// TIA Portal project "XSFW_TIA31001_B0_V15.1" (V15.1) (continued)
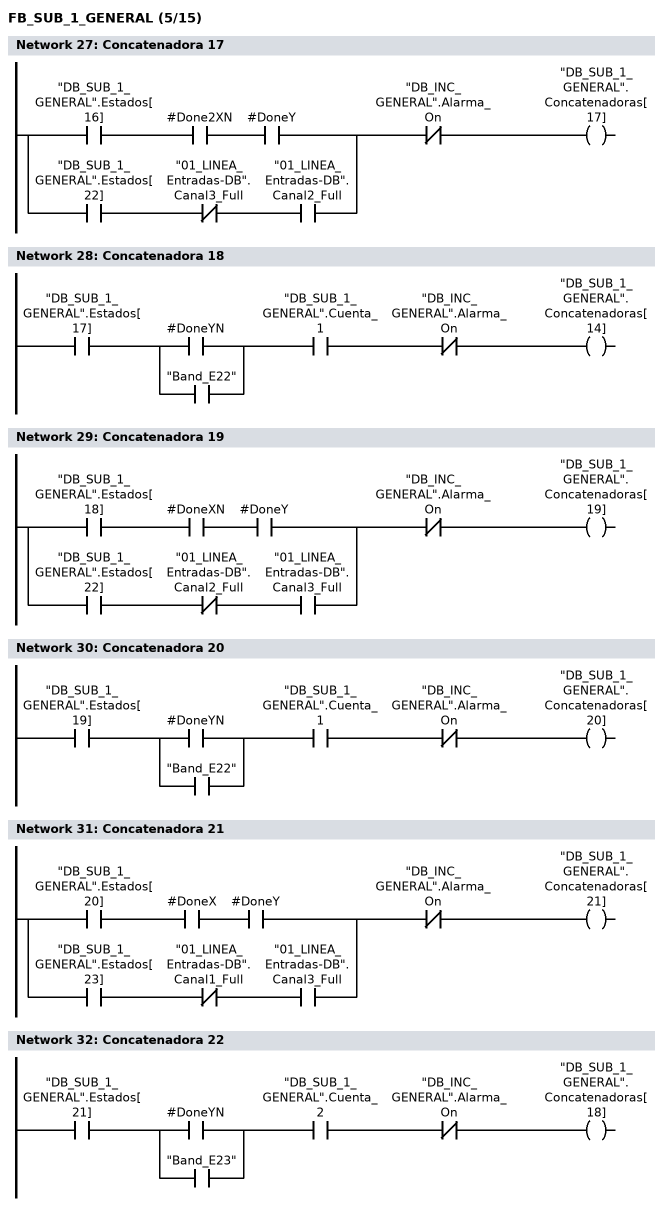
   RUNG wire#powerrail
      Contact( "DB_SUB_1_GENERAL".Estados[16] )
      Contact( #Done2XN )
      Contact( #DoneY )
      wire#w1
      I_Contact( "DB_INC_GENERAL".Alarma_On )
      Coil( "DB_SUB_1_GENERAL".Concatenadoras[17] )
   END_RUNG
   RUNG wire#powerrail
      Contact( "DB_SUB_1_GENERAL".Estados[22] )
      I_Contact( "01_LINEA_Entradas-DB".Canal3_Full )
      Contact( "01_LINEA_Entradas-DB".Canal2_Full )
   END_RUNG wire#w1
   // the same network as SCL:
   "DB_SUB_1_GENERAL".Concatenadoras[17] := (("DB_SUB_1_GENERAL".Estados[16] AND #Done2XN AND #DoneY) OR ("DB_SUB_1_GENERAL".Estados[22] AND NOT "01_LINEA_Entradas-DB".Canal3_Full AND "01_LINEA_Entradas-DB".Canal2_Full)) AND NOT "DB_INC_GENERAL".Alarma_On;
END_REGION

REGION Network 28: Concatenadora 18
   RUNG wire#powerrail
      Contact( "DB_SUB_1_GENERAL".Estados[17] )
      wire#w1
      Contact( #DoneYN )
      wire#w2
      Contact( "DB_SUB_1_GENERAL".Cuenta_1 )
      I_Contact( "DB_INC_GENERAL".Alarma_On )
      Coil( "DB_SUB_1_GENERAL".Concatenadoras[14] )
   END_RUNG
   RUNG wire#w1
      Contact( "Band_E22" )
   END_RUNG wire#w2
   // the same network as SCL:
   "DB_SUB_1_GENERAL".Concatenadoras[14] := "DB_SUB_1_GENERAL".Estados[17] AND (#DoneYN OR "Band_E22") AND "DB_SUB_1_GENERAL".Cuenta_1 AND NOT "DB_INC_GENERAL".Alarma_On;
END_REGION

REGION Network 29: Concatenadora 19
   RUNG wire#powerrail
      Contact( "DB_SUB_1_GENERAL".Estados[18] )
      Contact( #DoneXN )
      Contact( #DoneY )
      wire#w1
      I_Contact( "DB_INC_GENERAL".Alarma_On )
      Coil( "DB_SUB_1_GENERAL".Concatenadoras[19] )
   END_RUNG
   RUNG wire#powerrail
      Contact( "DB_SUB_1_GENERAL".Estados[22] )
      I_Contact( "01_LINEA_Entradas-DB".Canal2_Full )
      Contact( "01_LINEA_Entradas-DB".Canal3_Full )
   END_RUNG wire#w1
   // the same network as SCL:
   "DB_SUB_1_GENERAL".Concatenadoras[19] := (("DB_SUB_1_GENERAL".Estados[18] AND #DoneXN AND #DoneY) OR ("DB_SUB_1_GENERAL".Estados[22] AND NOT "01_LINEA_Entradas-DB".Canal2_Full AND "01_LINEA_Entradas-DB".Canal3_Full)) AND NOT "DB_INC_GENERAL".Alarma_On;
END_REGION

REGION Network 30: Concatenadora 20
   RUNG wire#powerrail
      Contact( "DB_SUB_1_GENERAL".Estados[19] )
      wire#w1
      Contact( #DoneYN )
      wire#w2
      Contact( "DB_SUB_1_GENERAL".Cuenta_1 )
      I_Contact( "DB_INC_GENERAL".Alarma_On )
      Coil( "DB_SUB_1_GENERAL".Concatenadoras[20] )
   END_RUNG
   RUNG wire#w1
      Contact( "Band_E22" )
   END_RUNG wire#w2
   // the same network as SCL:
   "DB_SUB_1_GENERAL".Concatenadoras[20] := "DB_SUB_1_GENERAL".Estados[19] AND (#DoneYN OR "Band_E22") AND "DB_SUB_1_GENERAL".Cuenta_1 AND NOT "DB_INC_GENERAL".Alarma_On;
END_REGION

REGION Network 31: Concatenadora 21
   RUNG wire#powerrail
      Contact( "DB_SUB_1_GENERAL".Estados[20] )
      Contact( #DoneX )
      Contact( #DoneY )
      wire#w1
      I_Contact( "DB_INC_GENERAL".Alarma_On )
      Coil( "DB_SUB_1_GENERAL".Concatenadoras[21] )
   END_RUNG
   RUNG wire#powerrail
      Contact( "DB_SUB_1_GENERAL".Estados[23] )
      I_Contact( "01_LINEA_Entradas-DB".Canal1_Full )
      Contact( "01_LINEA_Entradas-DB".Canal3_Full )
   END_RUNG wire#w1
   // the same network as SCL:
   "DB_SUB_1_GENERAL".Concatenadoras[21] := (("DB_SUB_1_GENERAL".Estados[20] AND #DoneX AND #DoneY) OR ("DB_SUB_1_GENERAL".Estados[23] AND NOT "01_LINEA_Entradas-DB".Canal1_Full AND "01_LINEA_Entradas-DB".Canal3_Full)) AND NOT "DB_INC_GENERAL".Alarma_On;
END_REGION

REGION Network 32: Concatenadora 22
   RUNG wire#powerrail
      Contact( "DB_SUB_1_GENERAL".Estados[21] )
      wire#w1
      Contact( #DoneYN )
      wire#w2
      Contact( "DB_SUB_1_GENERAL".Cuenta_2 )
      I_Contact( "DB_INC_GENERAL".Alarma_On )
      Coil( "DB_SUB_1_GENERAL".Concatenadoras[18] )
   END_RUNG
   RUNG wire#w1
      Contact( "Band_E23" )
   END_RUNG wire#w2
   // the same network as SCL:
   "DB_SUB_1_GENERAL".Concatenadoras[18] := "DB_SUB_1_GENERAL".Estados[21] AND (#DoneYN OR "Band_E23") AND "DB_SUB_1_GENERAL".Cuenta_2 AND NOT "DB_INC_GENERAL".Alarma_On;
END_REGION

REGION Network 33: Prioritaria 0
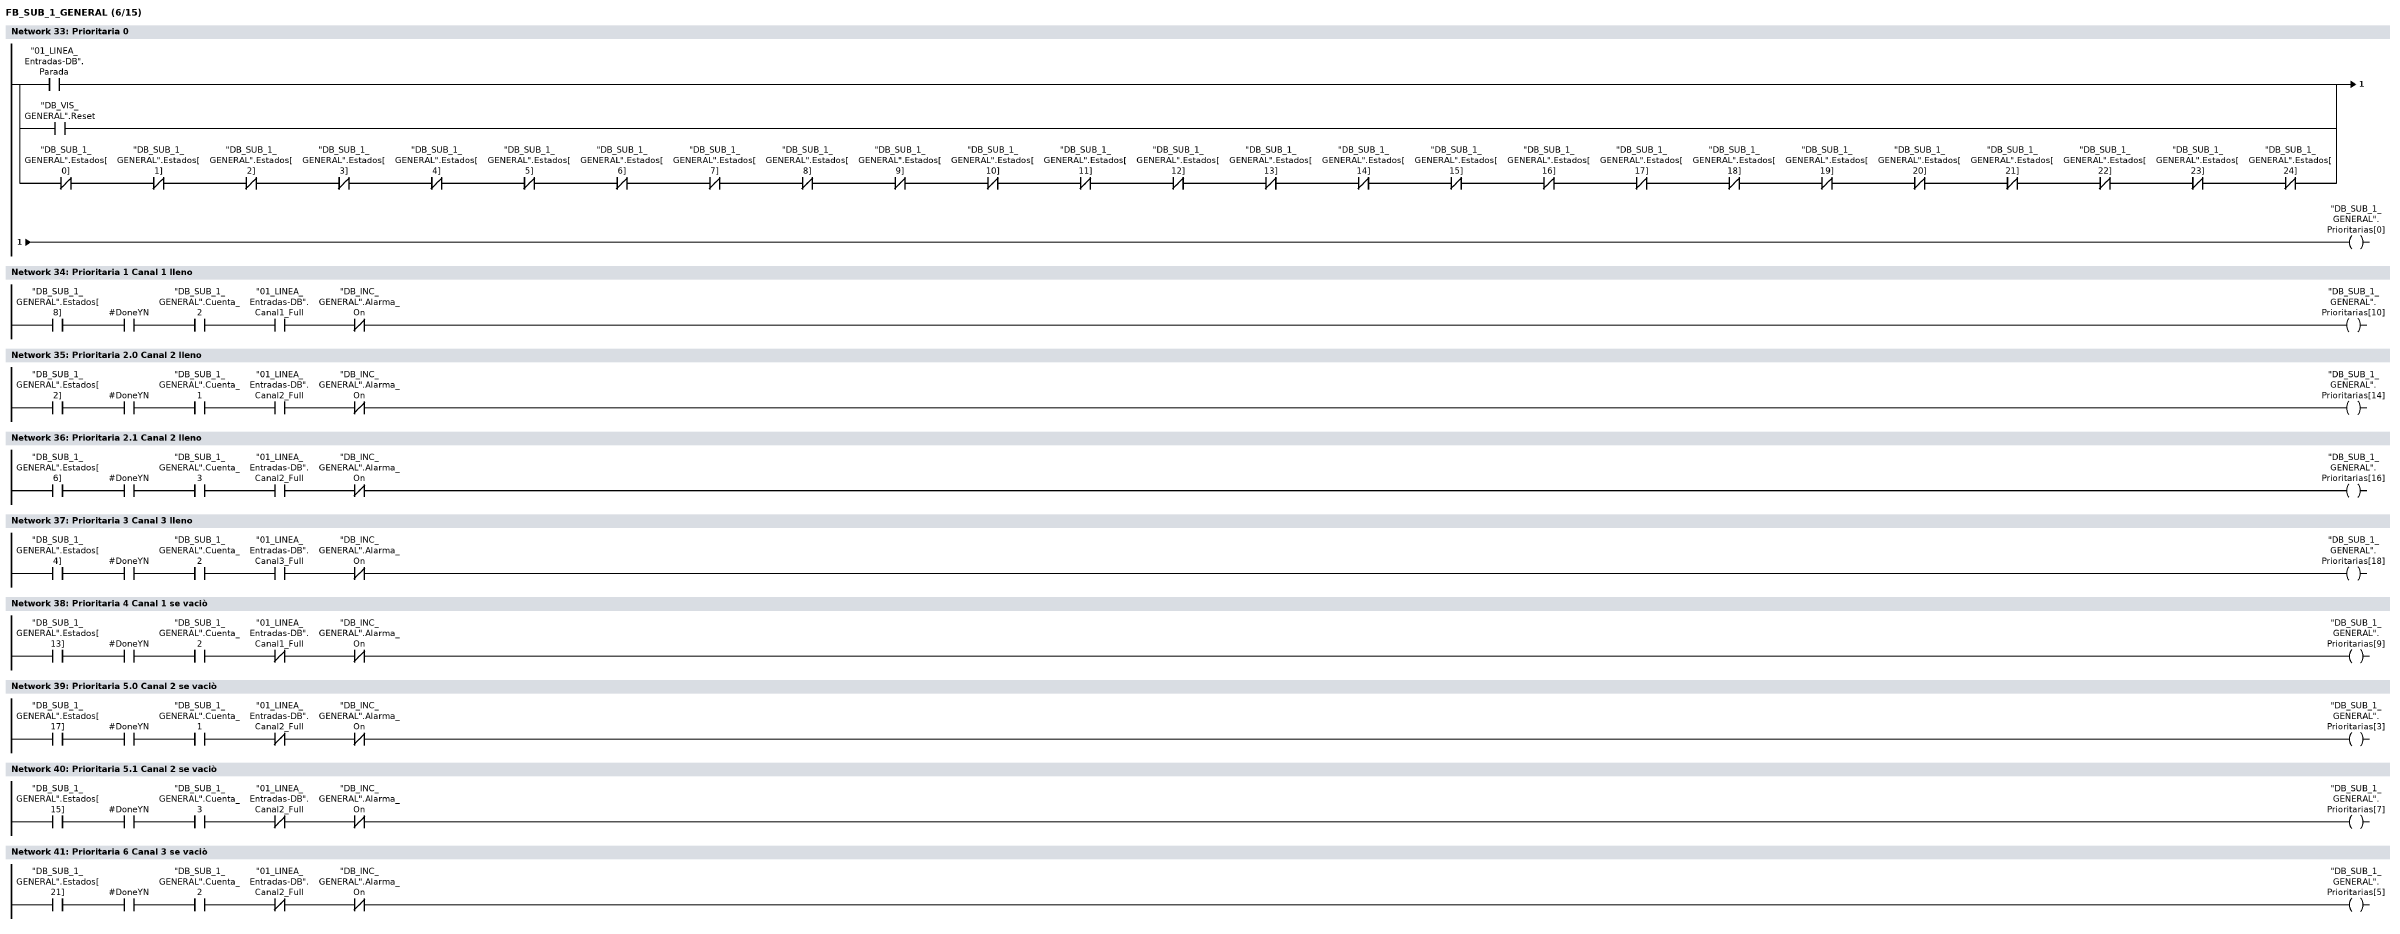
   RUNG wire#powerrail
      Contact( "01_LINEA_Entradas-DB".Parada )
      wire#w1
      Coil( "DB_SUB_1_GENERAL".Prioritarias[0] )
   END_RUNG
   RUNG wire#powerrail
      Contact( "DB_VIS_GENERAL".Reset )
   END_RUNG wire#w1
   RUNG wire#powerrail
      I_Contact( "DB_SUB_1_GENERAL".Estados[0] )
      I_Contact( "DB_SUB_1_GENERAL".Estados[1] )
      I_Contact( "DB_SUB_1_GENERAL".Estados[2] )
      I_Contact( "DB_SUB_1_GENERAL".Estados[3] )
      I_Contact( "DB_SUB_1_GENERAL".Estados[4] )
      I_Contact( "DB_SUB_1_GENERAL".Estados[5] )
      I_Contact( "DB_SUB_1_GENERAL".Estados[6] )
      I_Contact( "DB_SUB_1_GENERAL".Estados[7] )
      I_Contact( "DB_SUB_1_GENERAL".Estados[8] )
      I_Contact( "DB_SUB_1_GENERAL".Estados[9] )
      I_Contact( "DB_SUB_1_GENERAL".Estados[10] )
      I_Contact( "DB_SUB_1_GENERAL".Estados[11] )
      I_Contact( "DB_SUB_1_GENERAL".Estados[12] )
      I_Contact( "DB_SUB_1_GENERAL".Estados[13] )
      I_Contact( "DB_SUB_1_GENERAL".Estados[14] )
      I_Contact( "DB_SUB_1_GENERAL".Estados[15] )
      I_Contact( "DB_SUB_1_GENERAL".Estados[16] )
      I_Contact( "DB_SUB_1_GENERAL".Estados[17] )
      I_Contact( "DB_SUB_1_GENERAL".Estados[18] )
      I_Contact( "DB_SUB_1_GENERAL".Estados[19] )
      I_Contact( "DB_SUB_1_GENERAL".Estados[20] )
      I_Contact( "DB_SUB_1_GENERAL".Estados[21] )
      I_Contact( "DB_SUB_1_GENERAL".Estados[22] )
      I_Contact( "DB_SUB_1_GENERAL".Estados[23] )
      I_Contact( "DB_SUB_1_GENERAL".Estados[24] )
   END_RUNG wire#w1
   // the same network as SCL:
   "DB_SUB_1_GENERAL".Prioritarias[0] := "01_LINEA_Entradas-DB".Parada OR "DB_VIS_GENERAL".Reset OR (NOT "DB_SUB_1_GENERAL".Estados[0] AND NOT "DB_SUB_1_GENERAL".Estados[1] AND NOT "DB_SUB_1_GENERAL".Estados[2] AND NOT "DB_SUB_1_GENERAL".Estados[3] AND NOT "DB_SUB_1_GENERAL".Estados[4] AND NOT "DB_SUB_1_GENERAL".Estados[5] AND NOT "DB_SUB_1_GENERAL".Estados[6] AND NOT "DB_SUB_1_GENERAL".Estados[7] AND NOT "DB_SUB_1_GENERAL".Estados[8] AND NOT "DB_SUB_1_GENERAL".Estados[9] AND NOT "DB_SUB_1_GENERAL".Estados[10] AND NOT "DB_SUB_1_GENERAL".Estados[11] AND NOT "DB_SUB_1_GENERAL".Estados[12] AND NOT "DB_SUB_1_GENERAL".Estados[13] AND NOT "DB_SUB_1_GENERAL".Estados[14] AND NOT "DB_SUB_1_GENERAL".Estados[15] AND NOT "DB_SUB_1_GENERAL".Estados[16] AND NOT "DB_SUB_1_GENERAL".Estados[17] AND NOT "DB_SUB_1_GENERAL".Estados[18] AND NOT "DB_SUB_1_GENERAL".Estados[19] AND NOT "DB_SUB_1_GENERAL".Estados[20] AND NOT "DB_SUB_1_GENERAL".Estados[21] AND NOT "DB_SUB_1_GENERAL".Estados[22] AND NOT "DB_SUB_1_GENERAL".Estados[23] AND NOT "DB_SUB_1_GENERAL".Estados[24]);
END_REGION

REGION Network 34: Prioritaria 1 Canal 1 lleno
   RUNG wire#powerrail
      Contact( "DB_SUB_1_GENERAL".Estados[8] )
      Contact( #DoneYN )
      Contact( "DB_SUB_1_GENERAL".Cuenta_2 )
      Contact( "01_LINEA_Entradas-DB".Canal1_Full )
      I_Contact( "DB_INC_GENERAL".Alarma_On )
      Coil( "DB_SUB_1_GENERAL".Prioritarias[10] )
   END_RUNG
   // the same network as SCL:
   "DB_SUB_1_GENERAL".Prioritarias[10] := "DB_SUB_1_GENERAL".Estados[8] AND #DoneYN AND "DB_SUB_1_GENERAL".Cuenta_2 AND "01_LINEA_Entradas-DB".Canal1_Full AND NOT "DB_INC_GENERAL".Alarma_On;
END_REGION

REGION Network 35: Prioritaria 2.0 Canal 2 lleno
   RUNG wire#powerrail
      Contact( "DB_SUB_1_GENERAL".Estados[2] )
      Contact( #DoneYN )
      Contact( "DB_SUB_1_GENERAL".Cuenta_1 )
      Contact( "01_LINEA_Entradas-DB".Canal2_Full )
      I_Contact( "DB_INC_GENERAL".Alarma_On )
      Coil( "DB_SUB_1_GENERAL".Prioritarias[14] )
   END_RUNG
   // the same network as SCL:
   "DB_SUB_1_GENERAL".Prioritarias[14] := "DB_SUB_1_GENERAL".Estados[2] AND #DoneYN AND "DB_SUB_1_GENERAL".Cuenta_1 AND "01_LINEA_Entradas-DB".Canal2_Full AND NOT "DB_INC_GENERAL".Alarma_On;
END_REGION

REGION Network 36: Prioritaria 2.1 Canal 2 lleno
   RUNG wire#powerrail
      Contact( "DB_SUB_1_GENERAL".Estados[6] )
      Contact( #DoneYN )
      Contact( "DB_SUB_1_GENERAL".Cuenta_3 )
      Contact( "01_LINEA_Entradas-DB".Canal2_Full )
      I_Contact( "DB_INC_GENERAL".Alarma_On )
      Coil( "DB_SUB_1_GENERAL".Prioritarias[16] )
   END_RUNG
   // the same network as SCL:
   "DB_SUB_1_GENERAL".Prioritarias[16] := "DB_SUB_1_GENERAL".Estados[6] AND #DoneYN AND "DB_SUB_1_GENERAL".Cuenta_3 AND "01_LINEA_Entradas-DB".Canal2_Full AND NOT "DB_INC_GENERAL".Alarma_On;
END_REGION

REGION Network 37: Prioritaria 3 Canal 3 lleno
   RUNG wire#powerrail
      Contact( "DB_SUB_1_GENERAL".Estados[4] )
      Contact( #DoneYN )
      Contact( "DB_SUB_1_GENERAL".Cuenta_2 )
      Contact( "01_LINEA_Entradas-DB".Canal3_Full )
      I_Contact( "DB_INC_GENERAL".Alarma_On )
      Coil( "DB_SUB_1_GENERAL".Prioritarias[18] )
   END_RUNG
   // the same network as SCL:
   "DB_SUB_1_GENERAL".Prioritarias[18] := "DB_SUB_1_GENERAL".Estados[4] AND #DoneYN AND "DB_SUB_1_GENERAL".Cuenta_2 AND "01_LINEA_Entradas-DB".Canal3_Full AND NOT "DB_INC_GENERAL".Alarma_On;
END_REGION

REGION Network 38: Prioritaria 4 Canal 1 se vaciò
   RUNG wire#powerrail
      Contact( "DB_SUB_1_GENERAL".Estados[13] )
      Contact( #DoneYN )
      Contact( "DB_SUB_1_GENERAL".Cuenta_2 )
      I_Contact( "01_LINEA_Entradas-DB".Canal1_Full )
      I_Contact( "DB_INC_GENERAL".Alarma_On )
      Coil( "DB_SUB_1_GENERAL".Prioritarias[9] )
   END_RUNG
   // the same network as SCL:
   "DB_SUB_1_GENERAL".Prioritarias[9] := "DB_SUB_1_GENERAL".Estados[13] AND #DoneYN AND "DB_SUB_1_GENERAL".Cuenta_2 AND NOT "01_LINEA_Entradas-DB".Canal1_Full AND NOT "DB_INC_GENERAL".Alarma_On;
END_REGION

REGION Network 39: Prioritaria 5.0 Canal 2 se vaciò
   RUNG wire#powerrail
      Contact( "DB_SUB_1_GENERAL".Estados[17] )
      Contact( #DoneYN )
      Contact( "DB_SUB_1_GENERAL".Cuenta_1 )
      I_Contact( "01_LINEA_Entradas-DB".Canal2_Full )
      I_Contact( "DB_INC_GENERAL".Alarma_On )
      Coil( "DB_SUB_1_GENERAL".Prioritarias[3] )
   END_RUNG
   // the same network as SCL:
   "DB_SUB_1_GENERAL".Prioritarias[3] := "DB_SUB_1_GENERAL".Estados[17] AND #DoneYN AND "DB_SUB_1_GENERAL".Cuenta_1 AND NOT "01_LINEA_Entradas-DB".Canal2_Full AND NOT "DB_INC_GENERAL".Alarma_On;
END_REGION

REGION Network 40: Prioritaria 5.1 Canal 2 se vaciò
   RUNG wire#powerrail
      Contact( "DB_SUB_1_GENERAL".Estados[15] )
      Contact( #DoneYN )
      Contact( "DB_SUB_1_GENERAL".Cuenta_3 )
      I_Contact( "01_LINEA_Entradas-DB".Canal2_Full )
      I_Contact( "DB_INC_GENERAL".Alarma_On )
      Coil( "DB_SUB_1_GENERAL".Prioritarias[7] )
   END_RUNG
   // the same network as SCL:
   "DB_SUB_1_GENERAL".Prioritarias[7] := "DB_SUB_1_GENERAL".Estados[15] AND #DoneYN AND "DB_SUB_1_GENERAL".Cuenta_3 AND NOT "01_LINEA_Entradas-DB".Canal2_Full AND NOT "DB_INC_GENERAL".Alarma_On;
END_REGION

REGION Network 41: Prioritaria 6 Canal 3 se vaciò
   RUNG wire#powerrail
      Contact( "DB_SUB_1_GENERAL".Estados[21] )
      Contact( #DoneYN )
      Contact( "DB_SUB_1_GENERAL".Cuenta_2 )
      I_Contact( "01_LINEA_Entradas-DB".Canal2_Full )
      I_Contact( "DB_INC_GENERAL".Alarma_On )
      Coil( "DB_SUB_1_GENERAL".Prioritarias[5] )
   END_RUNG
   // the same network as SCL:
   "DB_SUB_1_GENERAL".Prioritarias[5] := "DB_SUB_1_GENERAL".Estados[21] AND #DoneYN AND "DB_SUB_1_GENERAL".Cuenta_2 AND NOT "01_LINEA_Entradas-DB".Canal2_Full AND NOT "DB_INC_GENERAL".Alarma_On;
END_REGION

REGION Network 42: Prioritaria 7 Canal 2 y 3 llenos
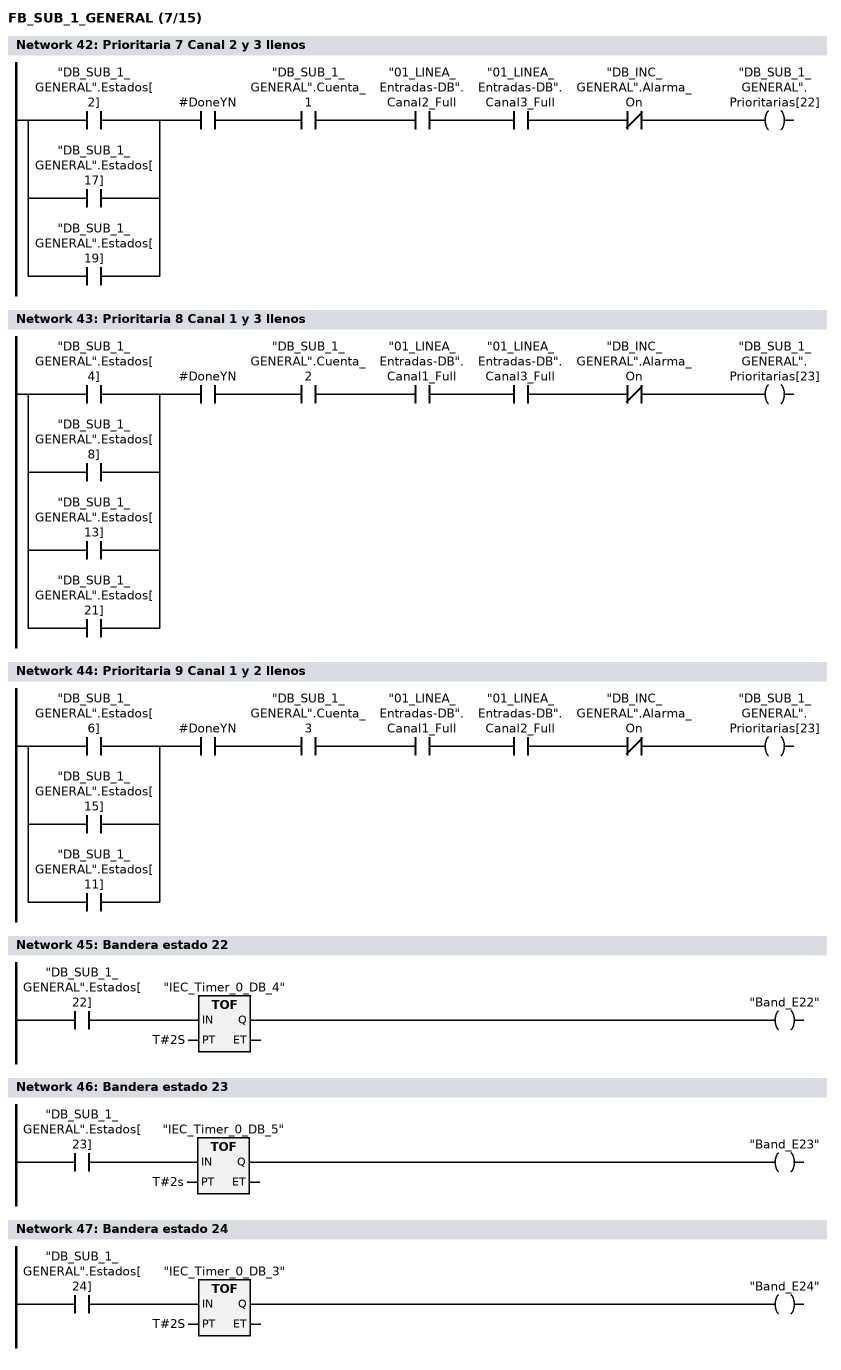
   RUNG wire#powerrail
      Contact( "DB_SUB_1_GENERAL".Estados[2] )
      wire#w1
      Contact( #DoneYN )
      Contact( "DB_SUB_1_GENERAL".Cuenta_1 )
      Contact( "01_LINEA_Entradas-DB".Canal2_Full )
      Contact( "01_LINEA_Entradas-DB".Canal3_Full )
      I_Contact( "DB_INC_GENERAL".Alarma_On )
      Coil( "DB_SUB_1_GENERAL".Prioritarias[22] )
   END_RUNG
   RUNG wire#powerrail
      Contact( "DB_SUB_1_GENERAL".Estados[17] )
   END_RUNG wire#w1
   RUNG wire#powerrail
      Contact( "DB_SUB_1_GENERAL".Estados[19] )
   END_RUNG wire#w1
   // the same network as SCL:
   "DB_SUB_1_GENERAL".Prioritarias[22] := ("DB_SUB_1_GENERAL".Estados[2] OR "DB_SUB_1_GENERAL".Estados[17] OR "DB_SUB_1_GENERAL".Estados[19]) AND #DoneYN AND "DB_SUB_1_GENERAL".Cuenta_1 AND "01_LINEA_Entradas-DB".Canal2_Full AND "01_LINEA_Entradas-DB".Canal3_Full AND NOT "DB_INC_GENERAL".Alarma_On;
END_REGION

REGION Network 43: Prioritaria 8 Canal 1 y 3 llenos
   RUNG wire#powerrail
      Contact( "DB_SUB_1_GENERAL".Estados[4] )
      wire#w1
      Contact( #DoneYN )
      Contact( "DB_SUB_1_GENERAL".Cuenta_2 )
      Contact( "01_LINEA_Entradas-DB".Canal1_Full )
      Contact( "01_LINEA_Entradas-DB".Canal3_Full )
      I_Contact( "DB_INC_GENERAL".Alarma_On )
      Coil( "DB_SUB_1_GENERAL".Prioritarias[23] )
   END_RUNG
   RUNG wire#powerrail
      Contact( "DB_SUB_1_GENERAL".Estados[8] )
   END_RUNG wire#w1
   RUNG wire#powerrail
      Contact( "DB_SUB_1_GENERAL".Estados[13] )
   END_RUNG wire#w1
   RUNG wire#powerrail
      Contact( "DB_SUB_1_GENERAL".Estados[21] )
   END_RUNG wire#w1
   // the same network as SCL:
   "DB_SUB_1_GENERAL".Prioritarias[23] := ("DB_SUB_1_GENERAL".Estados[4] OR "DB_SUB_1_GENERAL".Estados[8] OR "DB_SUB_1_GENERAL".Estados[13] OR "DB_SUB_1_GENERAL".Estados[21]) AND #DoneYN AND "DB_SUB_1_GENERAL".Cuenta_2 AND "01_LINEA_Entradas-DB".Canal1_Full AND "01_LINEA_Entradas-DB".Canal3_Full AND NOT "DB_INC_GENERAL".Alarma_On;
END_REGION

REGION Network 44: Prioritaria 9 Canal 1 y 2 llenos
   RUNG wire#powerrail
      Contact( "DB_SUB_1_GENERAL".Estados[6] )
      wire#w1
      Contact( #DoneYN )
      Contact( "DB_SUB_1_GENERAL".Cuenta_3 )
      Contact( "01_LINEA_Entradas-DB".Canal1_Full )
      Contact( "01_LINEA_Entradas-DB".Canal2_Full )
      I_Contact( "DB_INC_GENERAL".Alarma_On )
      Coil( "DB_SUB_1_GENERAL".Prioritarias[23] )
   END_RUNG
   RUNG wire#powerrail
      Contact( "DB_SUB_1_GENERAL".Estados[15] )
   END_RUNG wire#w1
   RUNG wire#powerrail
      Contact( "DB_SUB_1_GENERAL".Estados[11] )
   END_RUNG wire#w1
   // the same network as SCL:
   "DB_SUB_1_GENERAL".Prioritarias[23] := ("DB_SUB_1_GENERAL".Estados[6] OR "DB_SUB_1_GENERAL".Estados[15] OR "DB_SUB_1_GENERAL".Estados[11]) AND #DoneYN AND "DB_SUB_1_GENERAL".Cuenta_3 AND "01_LINEA_Entradas-DB".Canal1_Full AND "01_LINEA_Entradas-DB".Canal2_Full AND NOT "DB_INC_GENERAL".Alarma_On;
END_REGION

REGION Network 45: Bandera estado 22
   "IEC_Timer_0_DB_4".TOF(IN := "DB_SUB_1_GENERAL".Estados[22], PT := T#2S);
   "Band_E22" := "IEC_Timer_0_DB_4".Q;
END_REGION

REGION Network 46: Bandera estado 23
   "IEC_Timer_0_DB_5".TOF(IN := "DB_SUB_1_GENERAL".Estados[23], PT := T#2s);
   "Band_E23" := "IEC_Timer_0_DB_5".Q;
END_REGION

REGION Network 47: Bandera estado 24
   "IEC_Timer_0_DB_3".TOF(IN := "DB_SUB_1_GENERAL".Estados[24], PT := T#2S);
   "Band_E24" := "IEC_Timer_0_DB_3".Q;
END_REGION

REGION Network 48: BLOQUE MAQUINA ESTADO
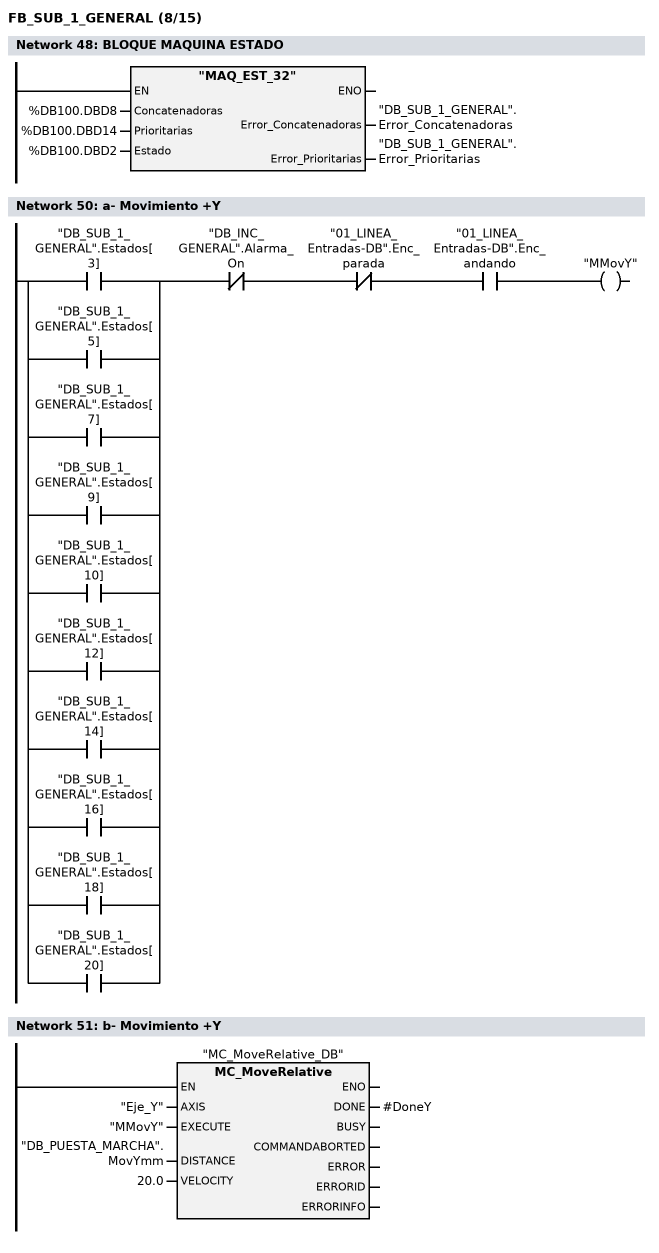
   RUNG wire#powerrail
      "MAQ_EST_32"(Concatenadoras := %DB100.DBD8, Prioritarias := %DB100.DBD14, Estado := %DB100.DBD2, Error_Concatenadoras => "DB_SUB_1_GENERAL".Error_Concatenadoras, Error_Prioritarias => "DB_SUB_1_GENERAL".Error_Prioritarias)
   END_RUNG
   // the same network as SCL:
   "MAQ_EST_32"(Concatenadoras := %DB100.DBD8,
                Prioritarias := %DB100.DBD14,
                Estado := %DB100.DBD2,
                Error_Concatenadoras => "DB_SUB_1_GENERAL".Error_Concatenadoras,
                Error_Prioritarias => "DB_SUB_1_GENERAL".Error_Prioritarias);
END_REGION

REGION Network 49: --------------ACCIONAMIENTOS----------------
END_REGION

REGION Network 50: a- Movimiento +Y
   RUNG wire#powerrail
      Contact( "DB_SUB_1_GENERAL".Estados[3] )
      wire#w1
      I_Contact( "DB_INC_GENERAL".Alarma_On )
      I_Contact( "01_LINEA_Entradas-DB".Enc_parada )
      Contact( "01_LINEA_Entradas-DB".Enc_andando )
      Coil( "MMovY" )
   END_RUNG
   RUNG wire#powerrail
      Contact( "DB_SUB_1_GENERAL".Estados[5] )
   END_RUNG wire#w1
   RUNG wire#powerrail
      Contact( "DB_SUB_1_GENERAL".Estados[7] )
   END_RUNG wire#w1
   RUNG wire#powerrail
      Contact( "DB_SUB_1_GENERAL".Estados[9] )
   END_RUNG wire#w1
   RUNG wire#powerrail
      Contact( "DB_SUB_1_GENERAL".Estados[10] )
   END_RUNG wire#w1
   RUNG wire#powerrail
      Contact( "DB_SUB_1_GENERAL".Estados[12] )
   END_RUNG wire#w1
   RUNG wire#powerrail
      Contact( "DB_SUB_1_GENERAL".Estados[14] )
   END_RUNG wire#w1
   RUNG wire#powerrail
      Contact( "DB_SUB_1_GENERAL".Estados[16] )
   END_RUNG wire#w1
   RUNG wire#powerrail
      Contact( "DB_SUB_1_GENERAL".Estados[18] )
   END_RUNG wire#w1
   RUNG wire#powerrail
      Contact( "DB_SUB_1_GENERAL".Estados[20] )
   END_RUNG wire#w1
   // the same network as SCL:
   "MMovY" := ("DB_SUB_1_GENERAL".Estados[3] OR "DB_SUB_1_GENERAL".Estados[5] OR "DB_SUB_1_GENERAL".Estados[7] OR "DB_SUB_1_GENERAL".Estados[9] OR "DB_SUB_1_GENERAL".Estados[10] OR "DB_SUB_1_GENERAL".Estados[12] OR "DB_SUB_1_GENERAL".Estados[14] OR "DB_SUB_1_GENERAL".Estados[16] OR "DB_SUB_1_GENERAL".Estados[18] OR "DB_SUB_1_GENERAL".Estados[20]) AND NOT "DB_INC_GENERAL".Alarma_On AND NOT "01_LINEA_Entradas-DB".Enc_parada AND "01_LINEA_Entradas-DB".Enc_andando;
END_REGION

REGION Network 51: b- Movimiento +Y
   "MC_MoveRelative_DB"(Axis := "Eje_Y",   // MC_MoveRelative
                        Execute := "MMovY",
                        Distance := "DB_PUESTA_MARCHA".MovYmm,
                        Velocity := 20.0,
                        Done => #DoneY);
END_REGION

REGION Network 52: a- Movimiento -Y
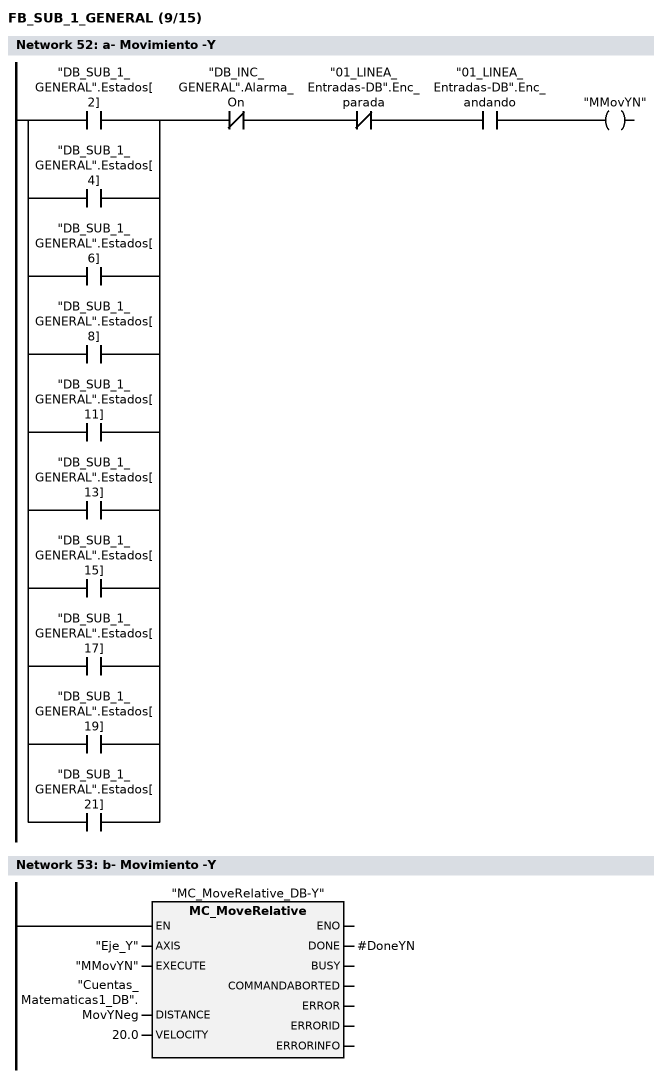
   RUNG wire#powerrail
      Contact( "DB_SUB_1_GENERAL".Estados[2] )
      wire#w1
      I_Contact( "DB_INC_GENERAL".Alarma_On )
      I_Contact( "01_LINEA_Entradas-DB".Enc_parada )
      Contact( "01_LINEA_Entradas-DB".Enc_andando )
      Coil( "MMovYN" )
   END_RUNG
   RUNG wire#powerrail
      Contact( "DB_SUB_1_GENERAL".Estados[4] )
   END_RUNG wire#w1
   RUNG wire#powerrail
      Contact( "DB_SUB_1_GENERAL".Estados[6] )
   END_RUNG wire#w1
   RUNG wire#powerrail
      Contact( "DB_SUB_1_GENERAL".Estados[8] )
   END_RUNG wire#w1
   RUNG wire#powerrail
      Contact( "DB_SUB_1_GENERAL".Estados[11] )
   END_RUNG wire#w1
   RUNG wire#powerrail
      Contact( "DB_SUB_1_GENERAL".Estados[13] )
   END_RUNG wire#w1
   RUNG wire#powerrail
      Contact( "DB_SUB_1_GENERAL".Estados[15] )
   END_RUNG wire#w1
   RUNG wire#powerrail
      Contact( "DB_SUB_1_GENERAL".Estados[17] )
   END_RUNG wire#w1
   RUNG wire#powerrail
      Contact( "DB_SUB_1_GENERAL".Estados[19] )
   END_RUNG wire#w1
   RUNG wire#powerrail
      Contact( "DB_SUB_1_GENERAL".Estados[21] )
   END_RUNG wire#w1
   // the same network as SCL:
   "MMovYN" := ("DB_SUB_1_GENERAL".Estados[2] OR "DB_SUB_1_GENERAL".Estados[4] OR "DB_SUB_1_GENERAL".Estados[6] OR "DB_SUB_1_GENERAL".Estados[8] OR "DB_SUB_1_GENERAL".Estados[11] OR "DB_SUB_1_GENERAL".Estados[13] OR "DB_SUB_1_GENERAL".Estados[15] OR "DB_SUB_1_GENERAL".Estados[17] OR "DB_SUB_1_GENERAL".Estados[19] OR "DB_SUB_1_GENERAL".Estados[21]) AND NOT "DB_INC_GENERAL".Alarma_On AND NOT "01_LINEA_Entradas-DB".Enc_parada AND "01_LINEA_Entradas-DB".Enc_andando;
END_REGION

REGION Network 53: b- Movimiento -Y
   "MC_MoveRelative_DB-Y"(Axis := "Eje_Y",   // MC_MoveRelative
                          Execute := "MMovYN",
                          Distance := "Cuentas_Matematicas1_DB".MovYNeg,
                          Velocity := 20.0,
                          Done => #DoneYN);
END_REGION

REGION Network 54: a- Movimiento +X
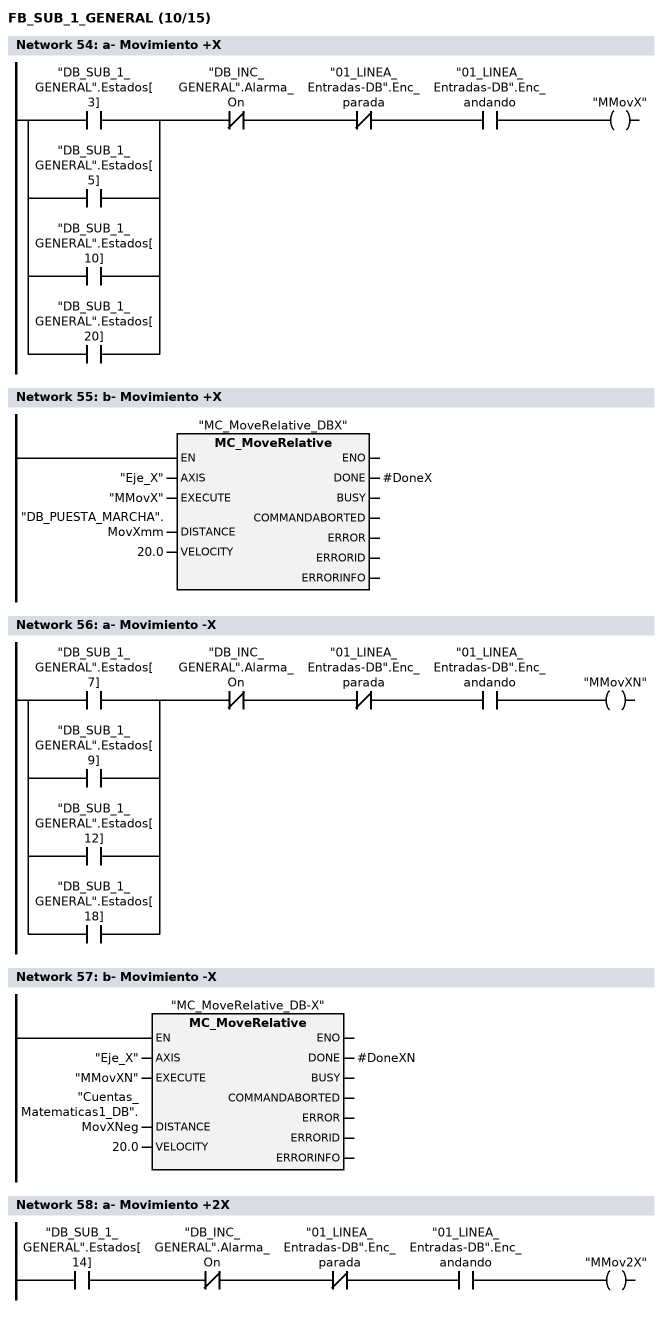
   RUNG wire#powerrail
      Contact( "DB_SUB_1_GENERAL".Estados[3] )
      wire#w1
      I_Contact( "DB_INC_GENERAL".Alarma_On )
      I_Contact( "01_LINEA_Entradas-DB".Enc_parada )
      Contact( "01_LINEA_Entradas-DB".Enc_andando )
      Coil( "MMovX" )
   END_RUNG
   RUNG wire#powerrail
      Contact( "DB_SUB_1_GENERAL".Estados[5] )
   END_RUNG wire#w1
   RUNG wire#powerrail
      Contact( "DB_SUB_1_GENERAL".Estados[10] )
   END_RUNG wire#w1
   RUNG wire#powerrail
      Contact( "DB_SUB_1_GENERAL".Estados[20] )
   END_RUNG wire#w1
   // the same network as SCL:
   "MMovX" := ("DB_SUB_1_GENERAL".Estados[3] OR "DB_SUB_1_GENERAL".Estados[5] OR "DB_SUB_1_GENERAL".Estados[10] OR "DB_SUB_1_GENERAL".Estados[20]) AND NOT "DB_INC_GENERAL".Alarma_On AND NOT "01_LINEA_Entradas-DB".Enc_parada AND "01_LINEA_Entradas-DB".Enc_andando;
END_REGION

REGION Network 55: b- Movimiento +X
   "MC_MoveRelative_DBX"(Axis := "Eje_X",   // MC_MoveRelative
                         Execute := "MMovX",
                         Distance := "DB_PUESTA_MARCHA".MovXmm,
                         Velocity := 20.0,
                         Done => #DoneX);
END_REGION

REGION Network 56: a- Movimiento -X
   RUNG wire#powerrail
      Contact( "DB_SUB_1_GENERAL".Estados[7] )
      wire#w1
      I_Contact( "DB_INC_GENERAL".Alarma_On )
      I_Contact( "01_LINEA_Entradas-DB".Enc_parada )
      Contact( "01_LINEA_Entradas-DB".Enc_andando )
      Coil( "MMovXN" )
   END_RUNG
   RUNG wire#powerrail
      Contact( "DB_SUB_1_GENERAL".Estados[9] )
   END_RUNG wire#w1
   RUNG wire#powerrail
      Contact( "DB_SUB_1_GENERAL".Estados[12] )
   END_RUNG wire#w1
   RUNG wire#powerrail
      Contact( "DB_SUB_1_GENERAL".Estados[18] )
   END_RUNG wire#w1
   // the same network as SCL:
   "MMovXN" := ("DB_SUB_1_GENERAL".Estados[7] OR "DB_SUB_1_GENERAL".Estados[9] OR "DB_SUB_1_GENERAL".Estados[12] OR "DB_SUB_1_GENERAL".Estados[18]) AND NOT "DB_INC_GENERAL".Alarma_On AND NOT "01_LINEA_Entradas-DB".Enc_parada AND "01_LINEA_Entradas-DB".Enc_andando;
END_REGION

REGION Network 57: b- Movimiento -X
   "MC_MoveRelative_DB-X"(Axis := "Eje_X",   // MC_MoveRelative
                          Execute := "MMovXN",
                          Distance := "Cuentas_Matematicas1_DB".MovXNeg,
                          Velocity := 20.0,
                          Done => #DoneXN);
END_REGION

REGION Network 58: a- Movimiento +2X
   RUNG wire#powerrail
      Contact( "DB_SUB_1_GENERAL".Estados[14] )
      I_Contact( "DB_INC_GENERAL".Alarma_On )
      I_Contact( "01_LINEA_Entradas-DB".Enc_parada )
      Contact( "01_LINEA_Entradas-DB".Enc_andando )
      Coil( "MMov2X" )
   END_RUNG
   // the same network as SCL:
   "MMov2X" := "DB_SUB_1_GENERAL".Estados[14] AND NOT "DB_INC_GENERAL".Alarma_On AND NOT "01_LINEA_Entradas-DB".Enc_parada AND "01_LINEA_Entradas-DB".Enc_andando;
END_REGION

REGION Network 59: b- Movimiento +2X
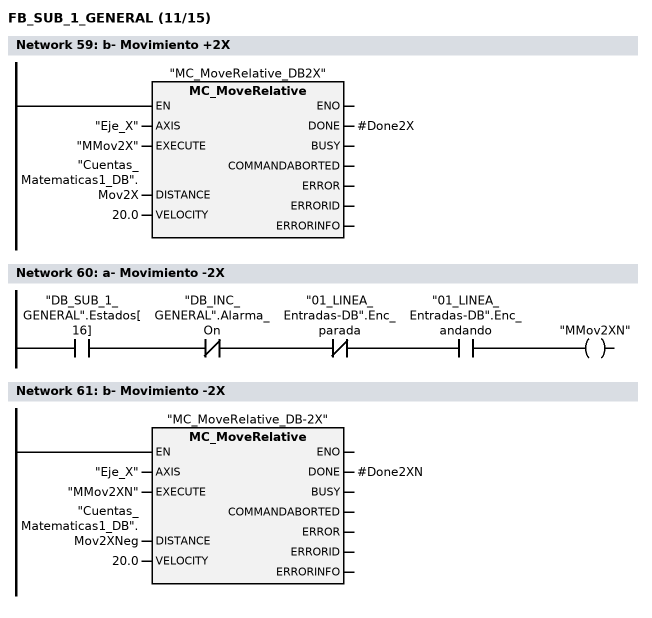
   "MC_MoveRelative_DB2X"(Axis := "Eje_X",   // MC_MoveRelative
                          Execute := "MMov2X",
                          Distance := "Cuentas_Matematicas1_DB".Mov2X,
                          Velocity := 20.0,
                          Done => #Done2X);
END_REGION

REGION Network 60: a- Movimiento -2X
   RUNG wire#powerrail
      Contact( "DB_SUB_1_GENERAL".Estados[16] )
      I_Contact( "DB_INC_GENERAL".Alarma_On )
      I_Contact( "01_LINEA_Entradas-DB".Enc_parada )
      Contact( "01_LINEA_Entradas-DB".Enc_andando )
      Coil( "MMov2XN" )
   END_RUNG
   // the same network as SCL:
   "MMov2XN" := "DB_SUB_1_GENERAL".Estados[16] AND NOT "DB_INC_GENERAL".Alarma_On AND NOT "01_LINEA_Entradas-DB".Enc_parada AND "01_LINEA_Entradas-DB".Enc_andando;
END_REGION

REGION Network 61: b- Movimiento -2X
   "MC_MoveRelative_DB-2X"(Axis := "Eje_X",   // MC_MoveRelative
                           Execute := "MMov2XN",
                           Distance := "Cuentas_Matematicas1_DB".Mov2XNeg,
                           Velocity := 20.0,
                           Done => #Done2XN);
END_REGION

REGION Network 62: Avance inverter